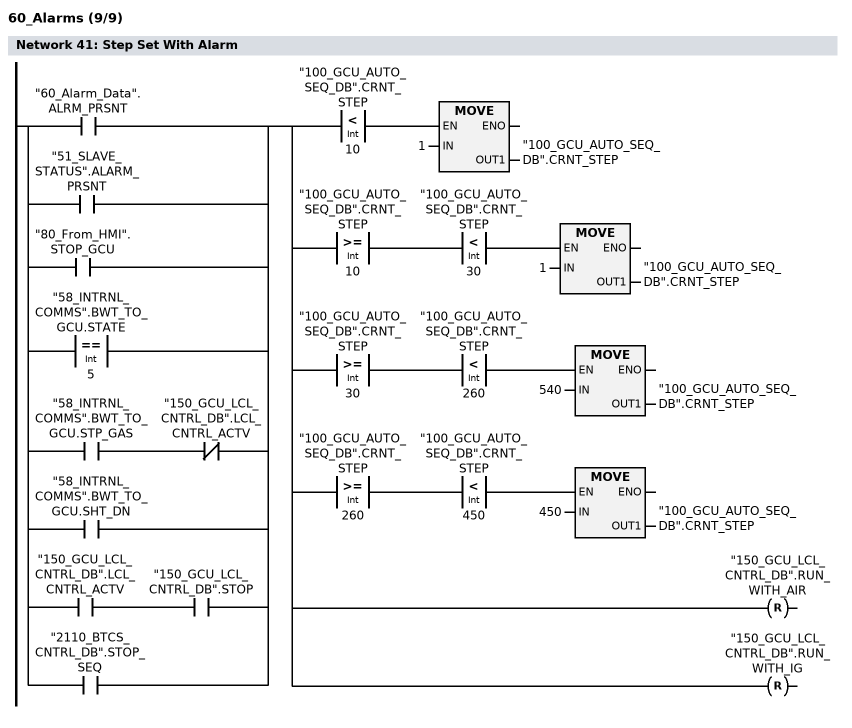
   RUNG wire#powerrail
      Contact( "60_Alarm_Data".ALRM_PRSNT )
      wire#w1
      { S7_Templates := "SrcType := Int" } LT_Contact(in1 := "100_GCU_AUTO_SEQ_DB".CRNT_STEP, in2 := 10)
      Move(in := 1, out1 => "100_GCU_AUTO_SEQ_DB".CRNT_STEP)
   END_RUNG
   RUNG wire#powerrail
      Contact( "51_SLAVE_STATUS".ALARM_PRSNT )
   END_RUNG wire#w1
   RUNG wire#powerrail
      Contact( "80_From_HMI".STOP_GCU )
   END_RUNG wire#w1
   RUNG wire#powerrail
      { S7_Templates := "SrcType := Int" } EQ_Contact(in1 := "58_INTRNL_COMMS".BWT_TO_GCU.STATE, in2 := 5)
   END_RUNG wire#w1
   RUNG wire#powerrail
      Contact( "58_INTRNL_COMMS".BWT_TO_GCU.STP_GAS )
      I_Contact( "150_GCU_LCL_CNTRL_DB".LCL_CNTRL_ACTV )
   END_RUNG wire#w1
   RUNG wire#powerrail
      Contact( "58_INTRNL_COMMS".BWT_TO_GCU.SHT_DN )
   END_RUNG wire#w1
   RUNG wire#powerrail
      Contact( "150_GCU_LCL_CNTRL_DB".LCL_CNTRL_ACTV )
      Contact( "150_GCU_LCL_CNTRL_DB".STOP )
   END_RUNG wire#w1
   RUNG wire#powerrail
      Contact( "2110_BTCS_CNTRL_DB".STOP_SEQ )
   END_RUNG wire#w1
   RUNG wire#w1
      { S7_Templates := "SrcType := Int" } GE_Contact(in1 := "100_GCU_AUTO_SEQ_DB".CRNT_STEP, in2 := 10)
      { S7_Templates := "SrcType := Int" } LT_Contact(in1 := "100_GCU_AUTO_SEQ_DB".CRNT_STEP, in2 := 30)
      Move(in := 1, out1 => "100_GCU_AUTO_SEQ_DB".CRNT_STEP)
   END_RUNG
   RUNG wire#w1
      { S7_Templates := "SrcType := Int" } GE_Contact(in1 := "100_GCU_AUTO_SEQ_DB".CRNT_STEP, in2 := 30)
      { S7_Templates := "SrcType := Int" } LT_Contact(in1 := "100_GCU_AUTO_SEQ_DB".CRNT_STEP, in2 := 260)
      Move(in := 540, out1 => "100_GCU_AUTO_SEQ_DB".CRNT_STEP)
   END_RUNG
   RUNG wire#w1
      { S7_Templates := "SrcType := Int" } GE_Contact(in1 := "100_GCU_AUTO_SEQ_DB".CRNT_STEP, in2 := 260)
      { S7_Templates := "SrcType := Int" } LT_Contact(in1 := "100_GCU_AUTO_SEQ_DB".CRNT_STEP, in2 := 450)
      Move(in := 450, out1 => "100_GCU_AUTO_SEQ_DB".CRNT_STEP)
   END_RUNG
   RUNG wire#w1
      R_Coil( "150_GCU_LCL_CNTRL_DB".RUN_WITH_AIR )
   END_RUNG
   RUNG wire#w1
      R_Coil( "150_GCU_LCL_CNTRL_DB".RUN_WITH_IG )
   END_RUNG
   // the same network as SCL:
   #_w1 := "60_Alarm_Data".ALRM_PRSNT OR "51_SLAVE_STATUS".ALARM_PRSNT OR "80_From_HMI".STOP_GCU OR ("58_INTRNL_COMMS".BWT_TO_GCU.STATE = 5) OR ("58_INTRNL_COMMS".BWT_TO_GCU.STP_GAS AND NOT "150_GCU_LCL_CNTRL_DB".LCL_CNTRL_ACTV) OR "58_INTRNL_COMMS".BWT_TO_GCU.SHT_DN OR ("150_GCU_LCL_CNTRL_DB".LCL_CNTRL_ACTV AND "150_GCU_LCL_CNTRL_DB".STOP) OR "2110_BTCS_CNTRL_DB".STOP_SEQ;
   IF #_w1 AND ("100_GCU_AUTO_SEQ_DB".CRNT_STEP < 10) THEN "100_GCU_AUTO_SEQ_DB".CRNT_STEP := 1; END_IF;
   IF #_w1 AND ("100_GCU_AUTO_SEQ_DB".CRNT_STEP >= 10) AND ("100_GCU_AUTO_SEQ_DB".CRNT_STEP < 30) THEN
       "100_GCU_AUTO_SEQ_DB".CRNT_STEP := 1;
   END_IF;
   IF #_w1 AND ("100_GCU_AUTO_SEQ_DB".CRNT_STEP >= 30) AND ("100_GCU_AUTO_SEQ_DB".CRNT_STEP < 260) THEN
       "100_GCU_AUTO_SEQ_DB".CRNT_STEP := 540;
   END_IF;
   IF #_w1 AND ("100_GCU_AUTO_SEQ_DB".CRNT_STEP >= 260) AND ("100_GCU_AUTO_SEQ_DB".CRNT_STEP < 450) THEN
       "100_GCU_AUTO_SEQ_DB".CRNT_STEP := 450;
   END_IF;
   IF #_w1 THEN
       "150_GCU_LCL_CNTRL_DB".RUN_WITH_AIR := FALSE;
       "150_GCU_LCL_CNTRL_DB".RUN_WITH_IG := FALSE;
   END_IF;
END_REGION
END_FUNCTION

FUNCTION "62_Warnings" : Void   // FC62, LAD
TITLE = Warning Processing
{ S7_Optimized_Access := 'TRUE' }
AUTHOR : JRS
VERSION : 0.1
// To warning conditions
   VAR_TEMP   // added for the SCL form of the ladder/FBD networks
      _w1 : Bool;
      _w2 : Bool;
   END_VAR
BEGIN

REGION Network 2: DB62 DBX2.0 =
   // GCU_WARNING_WORD_02_BIT_0
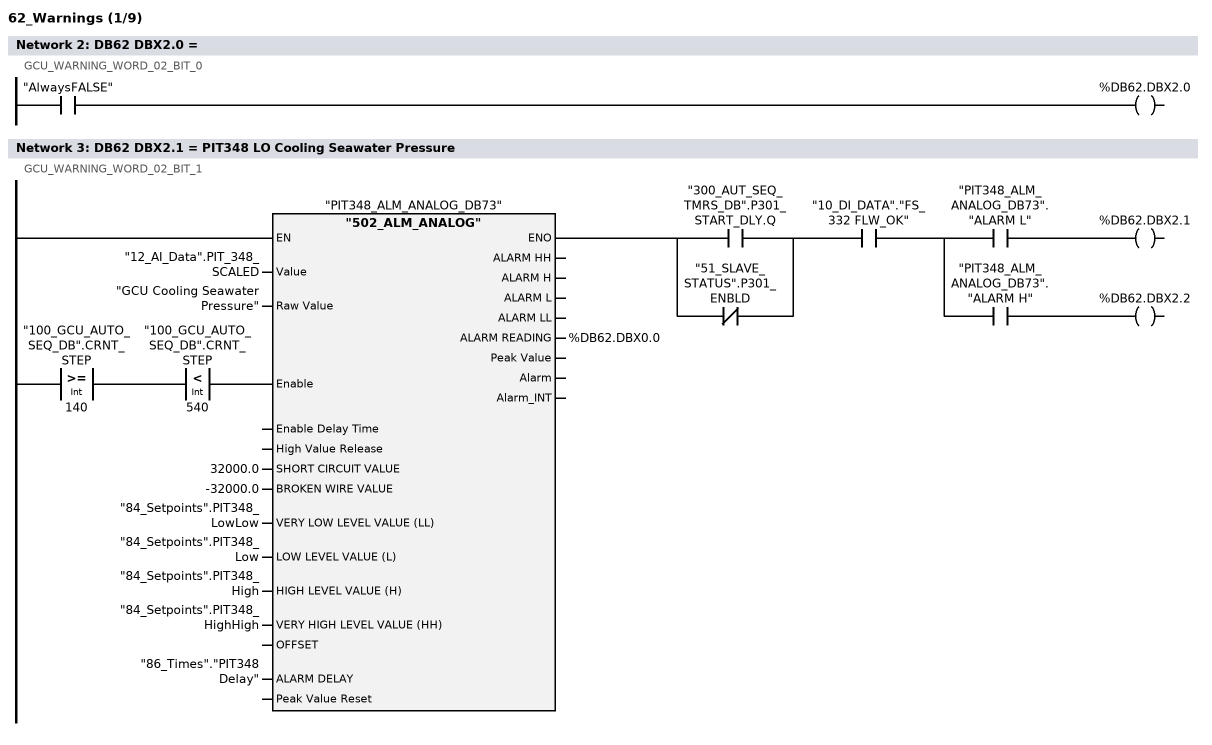
   RUNG wire#powerrail
      Contact( "AlwaysFALSE" )
      Coil( %DB62.DBX2.0 )
   END_RUNG
   // the same network as SCL:
   %DB62.DBX2.0 := "AlwaysFALSE";
END_REGION

REGION Network 3: DB62 DBX2.1 = PIT348 LO Cooling Seawater Pressure
   // GCU_WARNING_WORD_02_BIT_1
   RUNG wire#powerrail
      "PIT348_ALM_ANALOG_DB73"(Enable := wire#w1, Value := "12_AI_Data".PIT_348_SCALED, "Raw Value" := "GCU Cooling Seawater Pressure", "Enable Delay Time" :=, "High Value Release" :=, "SHORT CIRCUIT VALUE" := 32000.0, "BROKEN WIRE VALUE" := -32000.0, "VERY LOW LEVEL VALUE (LL)" := "84_Setpoints".PIT348_LowLow, "LOW LEVEL VALUE (L)" := "84_Setpoints".PIT348_Low, "HIGH LEVEL VALUE (H)" := "84_Setpoints".PIT348_High, "VERY HIGH LEVEL VALUE (HH)" := "84_Setpoints".PIT348_HighHigh, OFFSET :=, "ALARM DELAY" := "86_Times"."PIT348 Delay", "Peak Value Reset" :=, "ALARM HH" =>, "ALARM H" =>, "ALARM L" =>, "ALARM LL" =>, "ALARM READING" => %DB62.DBX0.0, "Peak Value" =>, Alarm =>, Alarm_INT =>)
      wire#w2
      Contact( "300_AUT_SEQ_TMRS_DB".P301_START_DLY.Q )
      wire#w3
      Contact( "10_DI_DATA"."FS_332 FLW_OK" )
      wire#w4
      Contact( "PIT348_ALM_ANALOG_DB73"."ALARM L" )
      Coil( %DB62.DBX2.1 )
   END_RUNG
   RUNG wire#powerrail
      { S7_Templates := "SrcType := Int" } GE_Contact(in1 := "100_GCU_AUTO_SEQ_DB".CRNT_STEP, in2 := 140)
      { S7_Templates := "SrcType := Int" } LT_Contact(in1 := "100_GCU_AUTO_SEQ_DB".CRNT_STEP, in2 := 540)
   END_RUNG wire#w1
   RUNG wire#w2
      I_Contact( "51_SLAVE_STATUS".P301_ENBLD )
   END_RUNG wire#w3
   RUNG wire#w4
      Contact( "PIT348_ALM_ANALOG_DB73"."ALARM H" )
      Coil( %DB62.DBX2.2 )
   END_RUNG
   // the same network as SCL:
   "PIT348_ALM_ANALOG_DB73"(Value := "12_AI_Data".PIT_348_SCALED,   // "502_ALM_ANALOG"
                           "Raw Value" := "GCU Cooling Seawater Pressure",
                           Enable := ("100_GCU_AUTO_SEQ_DB".CRNT_STEP >= 140) AND ("100_GCU_AUTO_SEQ_DB".CRNT_STEP < 540),
                           "SHORT CIRCUIT VALUE" := 32000.0,
                           "BROKEN WIRE VALUE" := -32000.0,
                           "VERY LOW LEVEL VALUE (LL)" := "84_Setpoints".PIT348_LowLow,
                           "LOW LEVEL VALUE (L)" := "84_Setpoints".PIT348_Low,
                           "HIGH LEVEL VALUE (H)" := "84_Setpoints".PIT348_High,
                           "VERY HIGH LEVEL VALUE (HH)" := "84_Setpoints".PIT348_HighHigh,
                           "ALARM DELAY" := "86_Times"."PIT348 Delay",
                           "ALARM READING" => %DB62.DBX0.0,
                           ENO => #_w1);
   #_w2 := #_w1 AND ("300_AUT_SEQ_TMRS_DB".P301_START_DLY.Q OR NOT "51_SLAVE_STATUS".P301_ENBLD) AND "10_DI_DATA"."FS_332 FLW_OK";
   %DB62.DBX2.1 := #_w2 AND "PIT348_ALM_ANALOG_DB73"."ALARM L";
   %DB62.DBX2.2 := #_w2 AND "PIT348_ALM_ANALOG_DB73"."ALARM H";
END_REGION

REGION Network 4: DB62 DBX2.3 = LIT304 GCU Tank Level HI / DB62 DBX2.4 = GCU Tank Level LO
   // GCU_WARNING_WORD_02_BIT_3
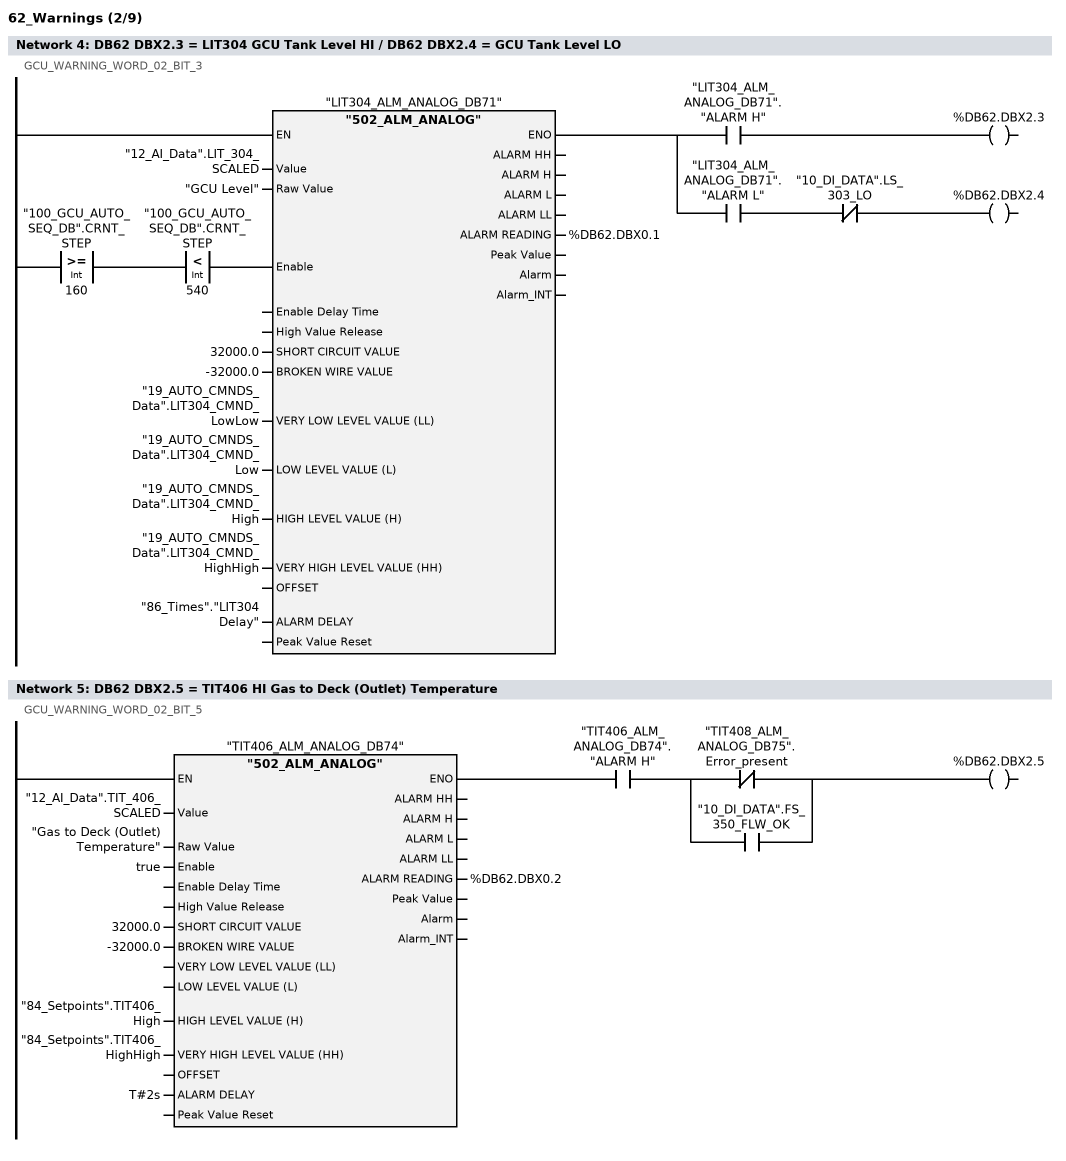
   RUNG wire#powerrail
      "LIT304_ALM_ANALOG_DB71"(Enable := wire#w1, Value := "12_AI_Data".LIT_304_SCALED, "Raw Value" := "GCU Level", "Enable Delay Time" :=, "High Value Release" :=, "SHORT CIRCUIT VALUE" := 32000.0, "BROKEN WIRE VALUE" := -32000.0, "VERY LOW LEVEL VALUE (LL)" := "19_AUTO_CMNDS_Data".LIT304_CMND_LowLow, "LOW LEVEL VALUE (L)" := "19_AUTO_CMNDS_Data".LIT304_CMND_Low, "HIGH LEVEL VALUE (H)" := "19_AUTO_CMNDS_Data".LIT304_CMND_High, "VERY HIGH LEVEL VALUE (HH)" := "19_AUTO_CMNDS_Data".LIT304_CMND_HighHigh, OFFSET :=, "ALARM DELAY" := "86_Times"."LIT304 Delay", "Peak Value Reset" :=, "ALARM HH" =>, "ALARM H" =>, "ALARM L" =>, "ALARM LL" =>, "ALARM READING" => %DB62.DBX0.1, "Peak Value" =>, Alarm =>, Alarm_INT =>)
      wire#w2
      Contact( "LIT304_ALM_ANALOG_DB71"."ALARM H" )
      Coil( %DB62.DBX2.3 )
   END_RUNG
   RUNG wire#powerrail
      { S7_Templates := "SrcType := Int" } GE_Contact(in1 := "100_GCU_AUTO_SEQ_DB".CRNT_STEP, in2 := 160)
      { S7_Templates := "SrcType := Int" } LT_Contact(in1 := "100_GCU_AUTO_SEQ_DB".CRNT_STEP, in2 := 540)
   END_RUNG wire#w1
   RUNG wire#w2
      Contact( "LIT304_ALM_ANALOG_DB71"."ALARM L" )
      I_Contact( "10_DI_DATA".LS_303_LO )
      Coil( %DB62.DBX2.4 )
   END_RUNG
   // the same network as SCL:
   "LIT304_ALM_ANALOG_DB71"(Value := "12_AI_Data".LIT_304_SCALED,   // "502_ALM_ANALOG"
                           "Raw Value" := "GCU Level",
                           Enable := ("100_GCU_AUTO_SEQ_DB".CRNT_STEP >= 160) AND ("100_GCU_AUTO_SEQ_DB".CRNT_STEP < 540),
                           "SHORT CIRCUIT VALUE" := 32000.0,
                           "BROKEN WIRE VALUE" := -32000.0,
                           "VERY LOW LEVEL VALUE (LL)" := "19_AUTO_CMNDS_Data".LIT304_CMND_LowLow,
                           "LOW LEVEL VALUE (L)" := "19_AUTO_CMNDS_Data".LIT304_CMND_Low,
                           "HIGH LEVEL VALUE (H)" := "19_AUTO_CMNDS_Data".LIT304_CMND_High,
                           "VERY HIGH LEVEL VALUE (HH)" := "19_AUTO_CMNDS_Data".LIT304_CMND_HighHigh,
                           "ALARM DELAY" := "86_Times"."LIT304 Delay",
                           "ALARM READING" => %DB62.DBX0.1,
                           ENO => #_w1);
   %DB62.DBX2.3 := #_w1 AND "LIT304_ALM_ANALOG_DB71"."ALARM H";
   %DB62.DBX2.4 := #_w1 AND "LIT304_ALM_ANALOG_DB71"."ALARM L" AND NOT "10_DI_DATA".LS_303_LO;
END_REGION

REGION Network 5: DB62 DBX2.5 = TIT406 HI Gas to Deck (Outlet) Temperature
   // GCU_WARNING_WORD_02_BIT_5
   RUNG wire#powerrail
      "TIT406_ALM_ANALOG_DB74"(Value := "12_AI_Data".TIT_406_SCALED, "Raw Value" := "Gas to Deck (Outlet) Temperature", Enable := true, "Enable Delay Time" :=, "High Value Release" :=, "SHORT CIRCUIT VALUE" := 32000.0, "BROKEN WIRE VALUE" := -32000.0, "VERY LOW LEVEL VALUE (LL)" :=, "LOW LEVEL VALUE (L)" :=, "HIGH LEVEL VALUE (H)" := "84_Setpoints".TIT406_High, "VERY HIGH LEVEL VALUE (HH)" := "84_Setpoints".TIT406_HighHigh, OFFSET :=, "ALARM DELAY" := T#2s, "Peak Value Reset" :=, "ALARM HH" =>, "ALARM H" =>, "ALARM L" =>, "ALARM LL" =>, "ALARM READING" => %DB62.DBX0.2, "Peak Value" =>, Alarm =>, Alarm_INT =>)
      Contact( "TIT406_ALM_ANALOG_DB74"."ALARM H" )
      wire#w1
      I_Contact( "TIT408_ALM_ANALOG_DB75".Error_present )
      wire#w2
      Coil( %DB62.DBX2.5 )
   END_RUNG
   RUNG wire#w1
      Contact( "10_DI_DATA".FS_350_FLW_OK )
   END_RUNG wire#w2
   // the same network as SCL:
   "TIT406_ALM_ANALOG_DB74"(Value := "12_AI_Data".TIT_406_SCALED,   // "502_ALM_ANALOG"
                           "Raw Value" := "Gas to Deck (Outlet) Temperature",
                           Enable := true,
                           "SHORT CIRCUIT VALUE" := 32000.0,
                           "BROKEN WIRE VALUE" := -32000.0,
                           "HIGH LEVEL VALUE (H)" := "84_Setpoints".TIT406_High,
                           "VERY HIGH LEVEL VALUE (HH)" := "84_Setpoints".TIT406_HighHigh,
                           "ALARM DELAY" := T#2s,
                           "ALARM READING" => %DB62.DBX0.2,
                           ENO => #_w1);
   %DB62.DBX2.5 := #_w1 AND "TIT406_ALM_ANALOG_DB74"."ALARM H" AND (NOT "TIT408_ALM_ANALOG_DB75".Error_present OR "10_DI_DATA".FS_350_FLW_OK);
END_REGION

REGION Network 6: DB62 DBX2.6 = TIT408 HI Fresh Water Cooling Temperature
   // GCU_WARNING_WORD_02_BIT_6
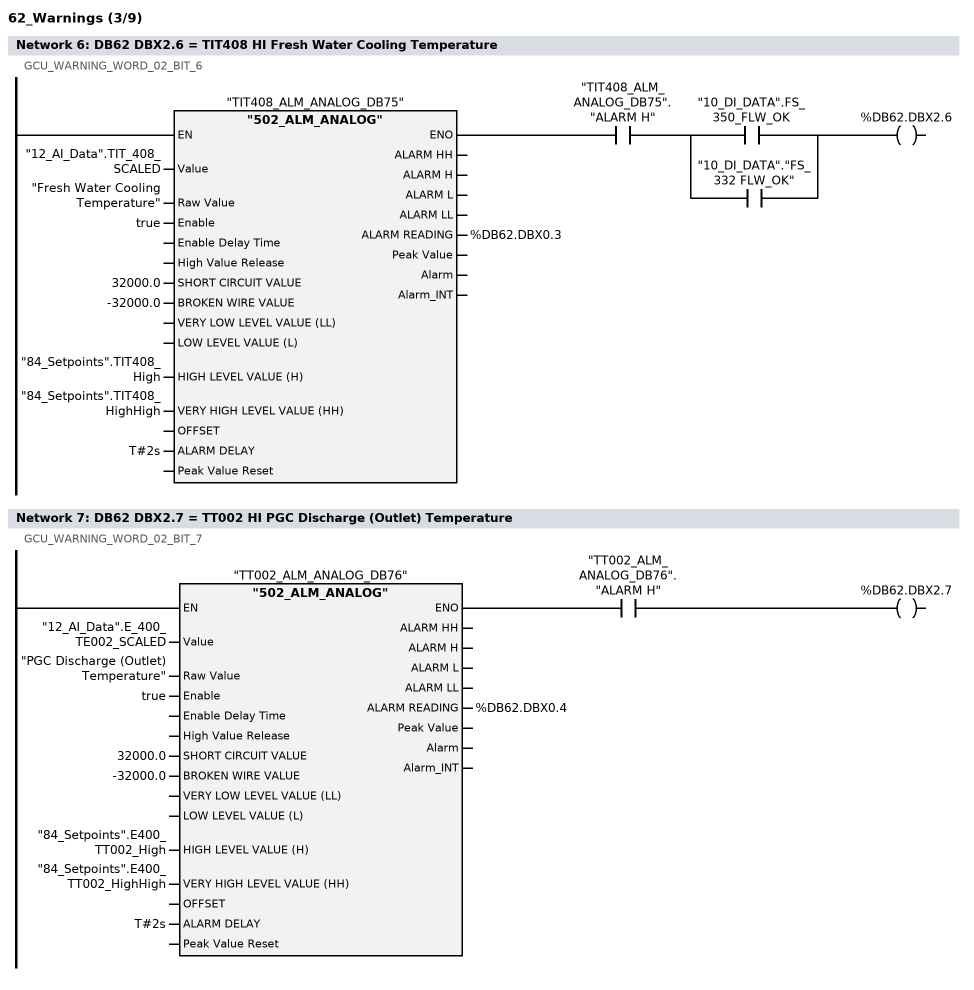
   RUNG wire#powerrail
      "TIT408_ALM_ANALOG_DB75"(Value := "12_AI_Data".TIT_408_SCALED, "Raw Value" := "Fresh Water Cooling Temperature", Enable := true, "Enable Delay Time" :=, "High Value Release" :=, "SHORT CIRCUIT VALUE" := 32000.0, "BROKEN WIRE VALUE" := -32000.0, "VERY LOW LEVEL VALUE (LL)" :=, "LOW LEVEL VALUE (L)" :=, "HIGH LEVEL VALUE (H)" := "84_Setpoints".TIT408_High, "VERY HIGH LEVEL VALUE (HH)" := "84_Setpoints".TIT408_HighHigh, OFFSET :=, "ALARM DELAY" := T#2s, "Peak Value Reset" :=, "ALARM HH" =>, "ALARM H" =>, "ALARM L" =>, "ALARM LL" =>, "ALARM READING" => %DB62.DBX0.3, "Peak Value" =>, Alarm =>, Alarm_INT =>)
      Contact( "TIT408_ALM_ANALOG_DB75"."ALARM H" )
      wire#w1
      Contact( "10_DI_DATA".FS_350_FLW_OK )
      wire#w2
      Coil( %DB62.DBX2.6 )
   END_RUNG
   RUNG wire#w1
      Contact( "10_DI_DATA"."FS_332 FLW_OK" )
   END_RUNG wire#w2
   // the same network as SCL:
   "TIT408_ALM_ANALOG_DB75"(Value := "12_AI_Data".TIT_408_SCALED,   // "502_ALM_ANALOG"
                           "Raw Value" := "Fresh Water Cooling Temperature",
                           Enable := true,
                           "SHORT CIRCUIT VALUE" := 32000.0,
                           "BROKEN WIRE VALUE" := -32000.0,
                           "HIGH LEVEL VALUE (H)" := "84_Setpoints".TIT408_High,
                           "VERY HIGH LEVEL VALUE (HH)" := "84_Setpoints".TIT408_HighHigh,
                           "ALARM DELAY" := T#2s,
                           "ALARM READING" => %DB62.DBX0.3,
                           ENO => #_w1);
   %DB62.DBX2.6 := #_w1 AND "TIT408_ALM_ANALOG_DB75"."ALARM H" AND ("10_DI_DATA".FS_350_FLW_OK OR "10_DI_DATA"."FS_332 FLW_OK");
END_REGION

REGION Network 7: DB62 DBX2.7 = TT002 HI PGC Discharge (Outlet) Temperature
   // GCU_WARNING_WORD_02_BIT_7
   RUNG wire#powerrail
      "TT002_ALM_ANALOG_DB76"(Value := "12_AI_Data".E_400_TE002_SCALED, "Raw Value" := "PGC Discharge (Outlet) Temperature", Enable := true, "Enable Delay Time" :=, "High Value Release" :=, "SHORT CIRCUIT VALUE" := 32000.0, "BROKEN WIRE VALUE" := -32000.0, "VERY LOW LEVEL VALUE (LL)" :=, "LOW LEVEL VALUE (L)" :=, "HIGH LEVEL VALUE (H)" := "84_Setpoints".E400_TT002_High, "VERY HIGH LEVEL VALUE (HH)" := "84_Setpoints".E400_TT002_HighHigh, OFFSET :=, "ALARM DELAY" := T#2s, "Peak Value Reset" :=, "ALARM HH" =>, "ALARM H" =>, "ALARM L" =>, "ALARM LL" =>, "ALARM READING" => %DB62.DBX0.4, "Peak Value" =>, Alarm =>, Alarm_INT =>)
      Contact( "TT002_ALM_ANALOG_DB76"."ALARM H" )
      Coil( %DB62.DBX2.7 )
   END_RUNG
   // the same network as SCL:
   "TT002_ALM_ANALOG_DB76"(Value := "12_AI_Data".E_400_TE002_SCALED,   // "502_ALM_ANALOG"
                           "Raw Value" := "PGC Discharge (Outlet) Temperature",
                           Enable := true,
                           "SHORT CIRCUIT VALUE" := 32000.0,
                           "BROKEN WIRE VALUE" := -32000.0,
                           "HIGH LEVEL VALUE (H)" := "84_Setpoints".E400_TT002_High,
                           "VERY HIGH LEVEL VALUE (HH)" := "84_Setpoints".E400_TT002_HighHigh,
                           "ALARM DELAY" := T#2s,
                           "ALARM READING" => %DB62.DBX0.4,
                           ENO => #_w1);
   %DB62.DBX2.7 := #_w1 AND "TT002_ALM_ANALOG_DB76"."ALARM H";
END_REGION

REGION Network 8: DB62 DBX3.0 = PT002 HI PGC Discharge (outlet) Pressure
   // GCU_WARNING_WORD_02_BIT_8
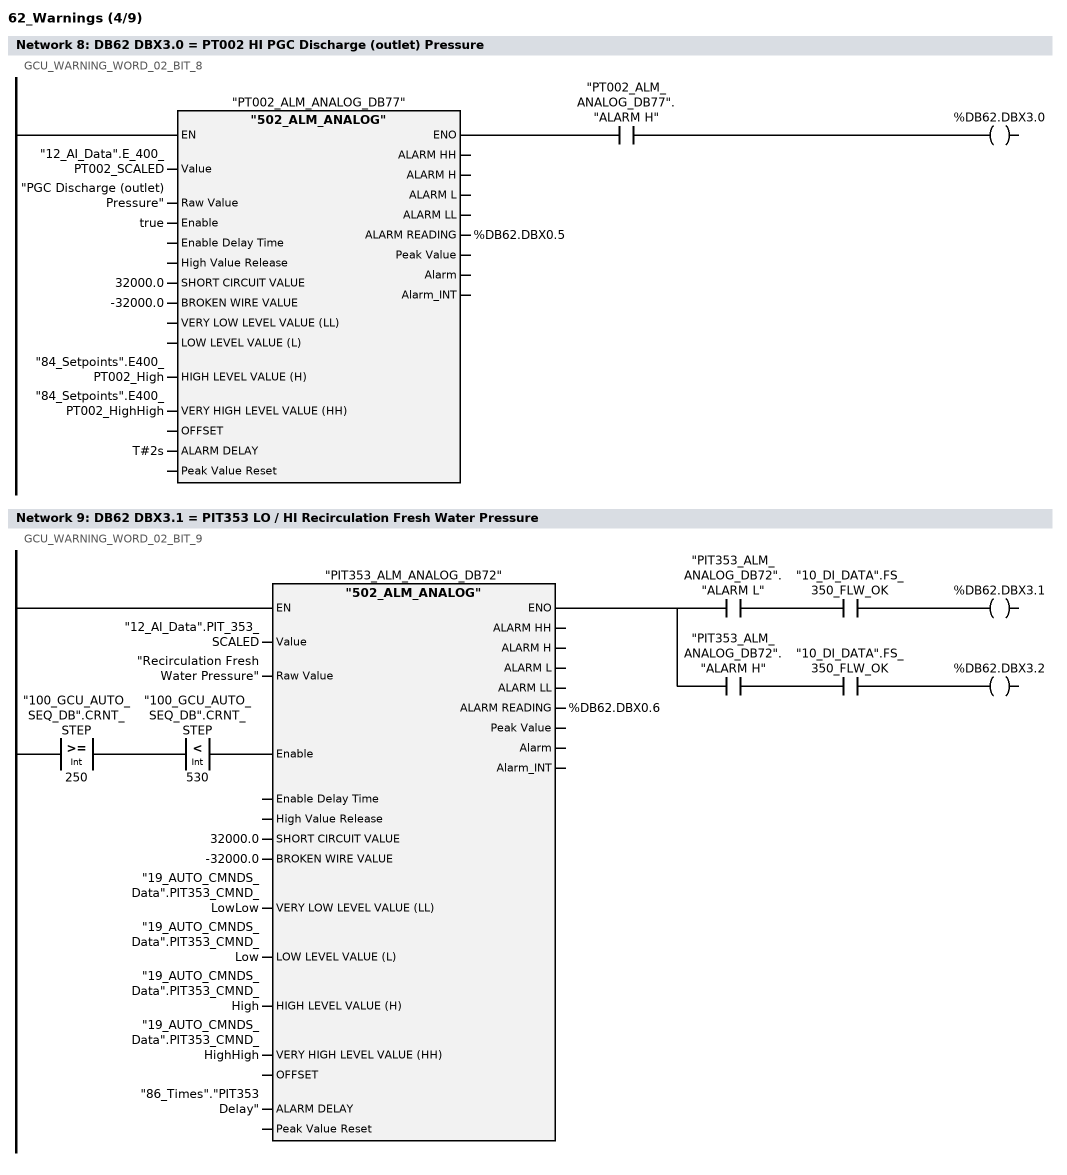
   RUNG wire#powerrail
      "PT002_ALM_ANALOG_DB77"(Value := "12_AI_Data".E_400_PT002_SCALED, "Raw Value" := "PGC Discharge (outlet) Pressure", Enable := true, "Enable Delay Time" :=, "High Value Release" :=, "SHORT CIRCUIT VALUE" := 32000.0, "BROKEN WIRE VALUE" := -32000.0, "VERY LOW LEVEL VALUE (LL)" :=, "LOW LEVEL VALUE (L)" :=, "HIGH LEVEL VALUE (H)" := "84_Setpoints".E400_PT002_High, "VERY HIGH LEVEL VALUE (HH)" := "84_Setpoints".E400_PT002_HighHigh, OFFSET :=, "ALARM DELAY" := T#2s, "Peak Value Reset" :=, "ALARM HH" =>, "ALARM H" =>, "ALARM L" =>, "ALARM LL" =>, "ALARM READING" => %DB62.DBX0.5, "Peak Value" =>, Alarm =>, Alarm_INT =>)
      Contact( "PT002_ALM_ANALOG_DB77"."ALARM H" )
      Coil( %DB62.DBX3.0 )
   END_RUNG
   // the same network as SCL:
   "PT002_ALM_ANALOG_DB77"(Value := "12_AI_Data".E_400_PT002_SCALED,   // "502_ALM_ANALOG"
                           "Raw Value" := "PGC Discharge (outlet) Pressure",
                           Enable := true,
                           "SHORT CIRCUIT VALUE" := 32000.0,
                           "BROKEN WIRE VALUE" := -32000.0,
                           "HIGH LEVEL VALUE (H)" := "84_Setpoints".E400_PT002_High,
                           "VERY HIGH LEVEL VALUE (HH)" := "84_Setpoints".E400_PT002_HighHigh,
                           "ALARM DELAY" := T#2s,
                           "ALARM READING" => %DB62.DBX0.5,
                           ENO => #_w1);
   %DB62.DBX3.0 := #_w1 AND "PT002_ALM_ANALOG_DB77"."ALARM H";
END_REGION

REGION Network 9: DB62 DBX3.1 = PIT353 LO / HI Recirculation Fresh Water Pressure
   // GCU_WARNING_WORD_02_BIT_9
   RUNG wire#powerrail
      "PIT353_ALM_ANALOG_DB72"(Enable := wire#w1, Value := "12_AI_Data".PIT_353_SCALED, "Raw Value" := "Recirculation Fresh Water Pressure", "Enable Delay Time" :=, "High Value Release" :=, "SHORT CIRCUIT VALUE" := 32000.0, "BROKEN WIRE VALUE" := -32000.0, "VERY LOW LEVEL VALUE (LL)" := "19_AUTO_CMNDS_Data".PIT353_CMND_LowLow, "LOW LEVEL VALUE (L)" := "19_AUTO_CMNDS_Data".PIT353_CMND_Low, "HIGH LEVEL VALUE (H)" := "19_AUTO_CMNDS_Data".PIT353_CMND_High, "VERY HIGH LEVEL VALUE (HH)" := "19_AUTO_CMNDS_Data".PIT353_CMND_HighHigh, OFFSET :=, "ALARM DELAY" := "86_Times"."PIT353 Delay", "Peak Value Reset" :=, "ALARM HH" =>, "ALARM H" =>, "ALARM L" =>, "ALARM LL" =>, "ALARM READING" => %DB62.DBX0.6, "Peak Value" =>, Alarm =>, Alarm_INT =>)
      wire#w2
      Contact( "PIT353_ALM_ANALOG_DB72"."ALARM L" )
      Contact( "10_DI_DATA".FS_350_FLW_OK )
      Coil( %DB62.DBX3.1 )
   END_RUNG
   RUNG wire#powerrail
      { S7_Templates := "SrcType := Int" } GE_Contact(in1 := "100_GCU_AUTO_SEQ_DB".CRNT_STEP, in2 := 250)
      { S7_Templates := "SrcType := Int" } LT_Contact(in1 := "100_GCU_AUTO_SEQ_DB".CRNT_STEP, in2 := 530)
   END_RUNG wire#w1
   RUNG wire#w2
      Contact( "PIT353_ALM_ANALOG_DB72"."ALARM H" )
      Contact( "10_DI_DATA".FS_350_FLW_OK )
      Coil( %DB62.DBX3.2 )
   END_RUNG
   // the same network as SCL:
   "PIT353_ALM_ANALOG_DB72"(Value := "12_AI_Data".PIT_353_SCALED,   // "502_ALM_ANALOG"
                           "Raw Value" := "Recirculation Fresh Water Pressure",
                           Enable := ("100_GCU_AUTO_SEQ_DB".CRNT_STEP >= 250) AND ("100_GCU_AUTO_SEQ_DB".CRNT_STEP < 530),
                           "SHORT CIRCUIT VALUE" := 32000.0,
                           "BROKEN WIRE VALUE" := -32000.0,
                           "VERY LOW LEVEL VALUE (LL)" := "19_AUTO_CMNDS_Data".PIT353_CMND_LowLow,
                           "LOW LEVEL VALUE (L)" := "19_AUTO_CMNDS_Data".PIT353_CMND_Low,
                           "HIGH LEVEL VALUE (H)" := "19_AUTO_CMNDS_Data".PIT353_CMND_High,
                           "VERY HIGH LEVEL VALUE (HH)" := "19_AUTO_CMNDS_Data".PIT353_CMND_HighHigh,
                           "ALARM DELAY" := "86_Times"."PIT353 Delay",
                           "ALARM READING" => %DB62.DBX0.6,
                           ENO => #_w1);
   %DB62.DBX3.1 := #_w1 AND "PIT353_ALM_ANALOG_DB72"."ALARM L" AND "10_DI_DATA".FS_350_FLW_OK;
   %DB62.DBX3.2 := #_w1 AND "PIT353_ALM_ANALOG_DB72"."ALARM H" AND "10_DI_DATA".FS_350_FLW_OK;
END_REGION

REGION Network 10: DB62 DBX3.3 = PIT416 LO Gas to Deck Pressure
   // GCU_WARNING_WORD_02_BIT_11      change from 450 to 520 as per Sequence sheet
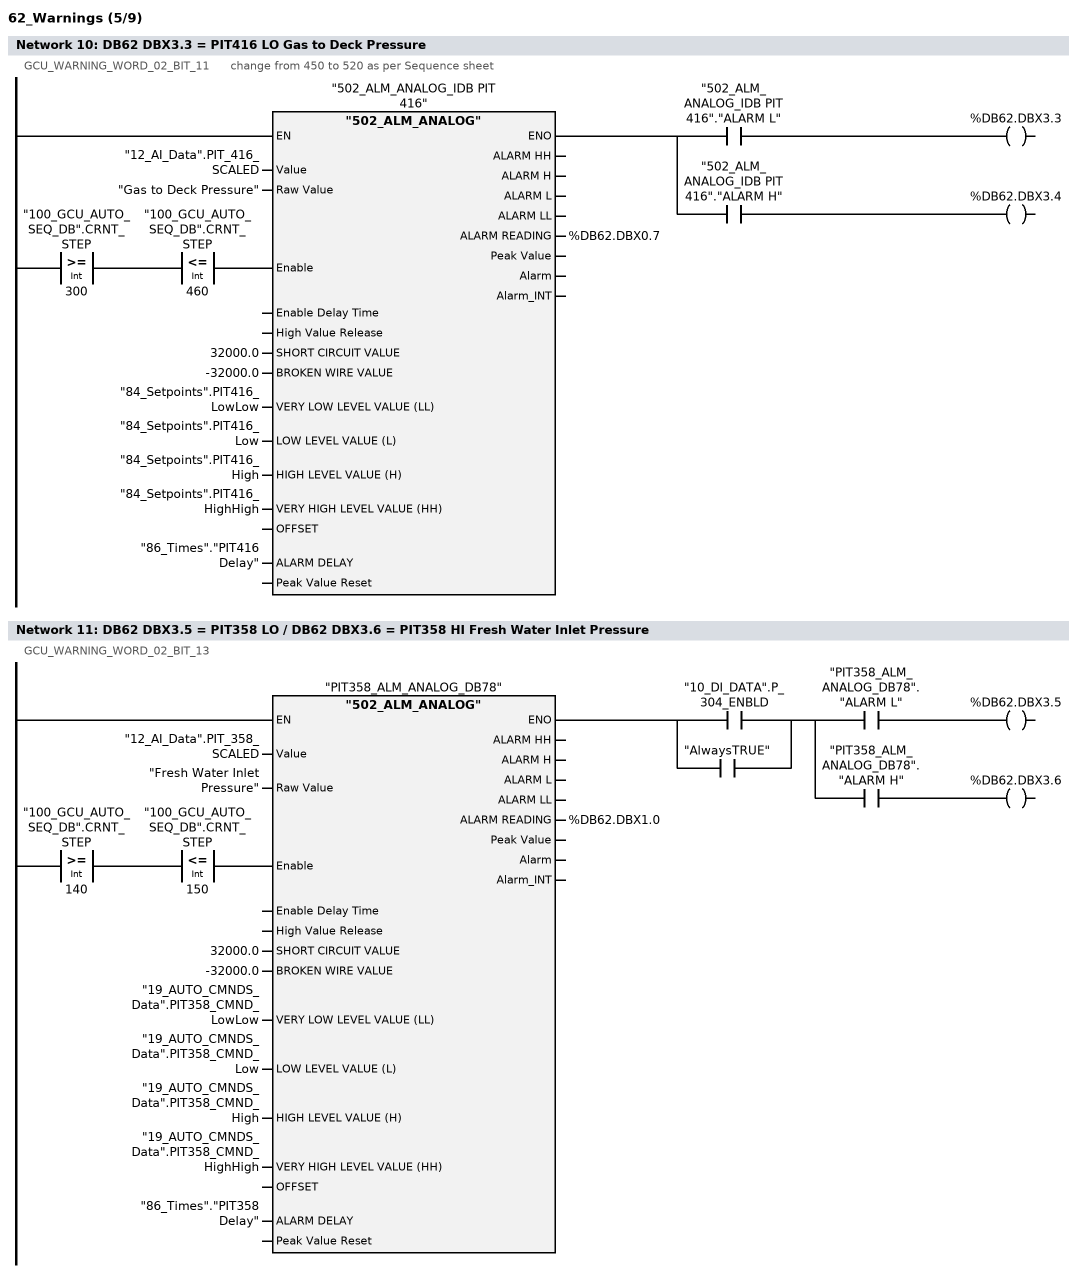
   RUNG wire#powerrail
      "502_ALM_ANALOG_IDB PIT 416"(Enable := wire#w1, Value := "12_AI_Data".PIT_416_SCALED, "Raw Value" := "Gas to Deck Pressure", "Enable Delay Time" :=, "High Value Release" :=, "SHORT CIRCUIT VALUE" := 32000.0, "BROKEN WIRE VALUE" := -32000.0, "VERY LOW LEVEL VALUE (LL)" := "84_Setpoints".PIT416_LowLow, "LOW LEVEL VALUE (L)" := "84_Setpoints".PIT416_Low, "HIGH LEVEL VALUE (H)" := "84_Setpoints".PIT416_High, "VERY HIGH LEVEL VALUE (HH)" := "84_Setpoints".PIT416_HighHigh, OFFSET :=, "ALARM DELAY" := "86_Times"."PIT416 Delay", "Peak Value Reset" :=, "ALARM HH" =>, "ALARM H" =>, "ALARM L" =>, "ALARM LL" =>, "ALARM READING" => %DB62.DBX0.7, "Peak Value" =>, Alarm =>, Alarm_INT =>)
      wire#w2
      Contact( "502_ALM_ANALOG_IDB PIT 416"."ALARM L" )
      Coil( %DB62.DBX3.3 )
   END_RUNG
   RUNG wire#powerrail
      { S7_Templates := "SrcType := Int" } GE_Contact(in1 := "100_GCU_AUTO_SEQ_DB".CRNT_STEP, in2 := 300)
      { S7_Templates := "SrcType := Int" } LE_Contact(in1 := "100_GCU_AUTO_SEQ_DB".CRNT_STEP, in2 := 460)
   END_RUNG wire#w1
   RUNG wire#w2
      Contact( "502_ALM_ANALOG_IDB PIT 416"."ALARM H" )
      Coil( %DB62.DBX3.4 )
   END_RUNG
   // the same network as SCL:
   "502_ALM_ANALOG_IDB PIT 416"(Value := "12_AI_Data".PIT_416_SCALED,   // "502_ALM_ANALOG"
                           "Raw Value" := "Gas to Deck Pressure",
                           Enable := ("100_GCU_AUTO_SEQ_DB".CRNT_STEP >= 300) AND ("100_GCU_AUTO_SEQ_DB".CRNT_STEP <= 460),
                           "SHORT CIRCUIT VALUE" := 32000.0,
                           "BROKEN WIRE VALUE" := -32000.0,
                           "VERY LOW LEVEL VALUE (LL)" := "84_Setpoints".PIT416_LowLow,
                           "LOW LEVEL VALUE (L)" := "84_Setpoints".PIT416_Low,
                           "HIGH LEVEL VALUE (H)" := "84_Setpoints".PIT416_High,
                           "VERY HIGH LEVEL VALUE (HH)" := "84_Setpoints".PIT416_HighHigh,
                           "ALARM DELAY" := "86_Times"."PIT416 Delay",
                           "ALARM READING" => %DB62.DBX0.7,
                           ENO => #_w1);
   %DB62.DBX3.3 := #_w1 AND "502_ALM_ANALOG_IDB PIT 416"."ALARM L";
   %DB62.DBX3.4 := #_w1 AND "502_ALM_ANALOG_IDB PIT 416"."ALARM H";
END_REGION
